// TIA Portal project "management parcare auto" (V17)

(* hardware
DEVICE "S7-1500/ET200MP station_1"  S7-1500 station
   slot 0: "Rail_0"  Rack  6ES7 590-1***0-0AA0
   slot 1: "PLC_1"  CPU 1511C-1 PN  6ES7 511-1CK01-0AB0  V2.5
      slot 3: "CPU display_1"  6ES7591-1AA00-0AA0
      slot 32768: "PROFINET interface_1"  X1
         slot 32769: "Port_1"  X1 P1
         slot 32770: "Port_2"  X1 P2
DEVICE "PC-System_1"  SIMATIC PC station
   slot 0: "SIMATIC PC station"  Rail  SIMATIC PC-Station  V1.0
      slot 125: "Stationmanager"  Station_Manager  V6.0.4
   slot 1: "HMI_RT_1"  WinCC RT Advanced  6AV2 104-0xxxx-xxxx  17.0.0.0
      slot 33792: "Computer interface"  Host interface
   slot 2: "CP 1628_1"  CP 1628  6GK1 162-8AA00  V8.2.2
DEVICE "HMI_1"  KTP700 Basic PN
   slot 0: "HMI_1"  KTP700 Basic PN  6AV2 123-2GB03-0AX0  15.1.0.0
   slot 1: "HMI_RT_2"  KTP700 Basic PN  6AV2 123-2GB03-0AX0  15.1.0.0
   slot 5: "HMI_1.IE_CP_1"  PROFINET Interface  15.0.1.0
      slot 1: "PROFINET Interface_1"  PROFINET Interface
         slot 1: "Port_1"  Port
*)

// ===== PLC "PLC_1"  CPU 1511C-1 PN =====

VAR_GLOBAL   // PLC tag table "Default tag table"
   "Exit barrier" AT %Q0.1 : Bool;
   "Entry barrier" AT %Q0.0 : Bool;
   "Entry sensor" AT %I0.0 : Bool;   // senzor bariera INTRARE
   "Exit sensor" AT %I1.0 : Bool;   // senzor barierea iesire
   "Parking lot 1 sensor" AT %I0.1 : Bool;   // senzor loc 1 (1-ocupat/ 0-liber)
   "Parking lot 2 sensor" AT %I0.2 : Bool;   // senzor loc 2
   "Parking lot 3 sensor" AT %I0.3 : Bool;
   "Parking lot 4 sensor" AT %I0.4 : Bool;
   "Parking lot 5 sensor" AT %I0.5 : Bool;
   "Parking lot 6 sensor" AT %I0.6 : Bool;
   "Parking lot 7 sensor" AT %I0.7 : Bool;
   "Parking lot 8 sensor" AT %I1.1 : Bool;
   "Parking lot 9 sensor" AT %I1.2 : Bool;
   "Parking lot 10 sensor" AT %I1.3 : Bool;
   "Number of cars" AT %MW20 : Int;   // nr de masini folosit la counter
   "System_Byte" AT %MB1 : Byte;
   "FirstScan" AT %M1.0 : Bool;
   "DiagStatusUpdate" AT %M1.1 : Bool;
   "AlwaysTRUE" AT %M1.2 : Bool;
   "AlwaysFALSE" AT %M1.3 : Bool;
   "Clock_Byte" AT %MB0 : Byte;
   "Clock_10Hz" AT %M0.0 : Bool;
   "Clock_5Hz" AT %M0.1 : Bool;
   "Clock_2.5Hz" AT %M0.2 : Bool;
   "Clock_2Hz" AT %M0.3 : Bool;
   "Clock_1.25Hz" AT %M0.4 : Bool;
   "Clock_1Hz" AT %M0.5 : Bool;
   "Clock_0.625Hz" AT %M0.6 : Bool;
   "Clock_0.5Hz" AT %M0.7 : Bool;
   "RdyToLog" AT %M2.0 : Bool;   // tagg folosit ca trigger pentru a rula vbScriptul
   "Tag5" AT %MW2 : Int;   // tagg folosit pentru counter pt animatie bariera intrare
   "Tag6" AT %MW4 : Int;   // tagg folosit pentru counter pt animatie bariera iesire
   "Tag_1" AT %M5.0 : Bool;
   "RdyToUpdate" AT %M6.0 : Bool;   // tagg folosit ca trigger pentru a rula vbSriptul de edit database
   "RdyToDelete" AT %M6.1 : Bool;   // tagg folosit ca trigger pentru a rula VbScriptul de stergere
   "Tag_2" AT %M6.2 : Bool;
   "Tag_3" AT %M6.3 : Bool;
   "Tag_4" AT %M6.4 : Bool;
   "Tag_5" AT %M6.5 : Bool;
   "Tag_6" AT %M6.6 : Bool;
   "Tag_7" AT %M6.7 : Bool;
   "Tag_8" AT %M5.1 : Bool;
   "Tag_9" AT %M5.2 : Bool;
   "Tag_10" AT %M5.3 : Bool;
   "Tag_11" AT %M5.4 : Bool;
   "Tag_12" AT %M7.0 : Bool;
   "Tag_13" AT %M7.1 : Bool;
   "Tag_14" AT %M7.2 : Bool;
   "Tag_15" AT %M7.3 : Bool;
   "Tag_16" AT %M7.4 : Bool;
   "Tag_17" AT %M7.5 : Bool;
   "Tag_18" AT %M7.6 : Bool;
   "Tag_19" AT %M7.7 : Bool;
   "Tag_20" AT %M8.0 : Bool;
   "Tag_21" AT %M8.1 : Bool;
END_VAR

// folder: DB's

DATA_BLOCK "02_DB_HMI_Buttons"   // DB2
{ S7_Optimized_Access := 'TRUE' }
VERSION : 0.1
   VAR
      pay : Bool;   // buton care simuleaza plata pentru a iesi din parcare
      "Parking lot 1" : Bool;   // buton in Hmi pentru a alege ce loc de parcare sa fie ocupat
      "Parking lot 2" : Bool;   // buton in Hmi pentru a alege ce loc de parcare sa fie ocupat
      "Parking lot 3" : Bool;   // buton in Hmi pentru a alege ce loc de parcare sa fie ocupat
      "Parking lot 4" : Bool;   // buton in Hmi pentru a alege ce loc de parcare sa fie ocupat
      "Parking lot 5" : Bool;   // buton in Hmi pentru a alege ce loc de parcare sa fie ocupat
      "Parking lot 6" : Bool;   // buton in Hmi pentru a alege ce loc de parcare sa fie ocupat
      "Parking lot 7" : Bool;   // buton in Hmi pentru a alege ce loc de parcare sa fie ocupat
      "Parking lot 8" : Bool;   // buton in Hmi pentru a alege ce loc de parcare sa fie ocupat
      "Parking lot 9" : Bool;   // buton in Hmi pentru a alege ce loc de parcare sa fie ocupat
      "Parking lot 10" : Bool;   // buton in Hmi pentru a alege ce loc de parcare sa fie ocupat
      "Entry button" : Bool;   // buton care simuleaza senzorul de intrare de la bariera
      "Exit button" : Bool;   // buton care simuleaza senzordul de iesire de la bariera
   END_VAR
   VAR RETAIN
      nrMasina_intrare : String;
   END_VAR
   VAR
      blank : String;
      nrMasina_iesire : String;
   END_VAR
BEGIN
END_DATA_BLOCK

DATA_BLOCK "04_DB_MarkersAuto"   // DB4
{ S7_Optimized_Access := 'TRUE' }
VERSION : 0.1
   VAR
      "car status_1" : Bool;
      "car status_2" : Bool;
      "car status_3" : Bool;
      "car status_4" : Bool;
      "car status_5" : Bool;
      "car status_6" : Bool;
      "car status_7" : Bool;
      "car status_8" : Bool;
      "car status_9" : Bool;
      "car status_10" : Bool;
      "remaining parking lots" : Int := 10;
      CarNumber : Int;   // dupa ce se introd un nr de masina, se face 1 , adica nr de masina a fost memorat
      "car status" : Bool;
      "Parking_lot_occupied 1" : Bool;   // locul a fost ocupat
      "Parking_lot_occupied 2" : Bool;
      "Parking_lot_occupied 3" : Bool;
      "Parking_lot_occupied 4" : Bool;
      "Parking_lot_occupied 5" : Bool;
      "Parking_lot_occupied 6" : Bool;
      "Parking_lot_occupied 7" : Bool;
      "Parking_lot_occupied 8" : Bool;
      "Parking_lot_occupied 9" : Bool;
      "Parking_lot_occupied 10" : Bool;
   END_VAR
BEGIN
END_DATA_BLOCK

DATA_BLOCK "05_DB_WinCC_buttons"   // DB5
{ S7_Optimized_Access := 'TRUE' }
VERSION : 0.1
   VAR
      loc_parcare_1 : Bool;   // buton de optiune pentru a alege locul de parcare 1
      loc_parcare_2 : Bool;   // -----//-------
      loc_parcare_3 : Bool;   // -----//-------
      loc_parcare_4 : Bool;   // -----//-------
      loc_parcare_5 : Bool;   // -----//-------
      loc_parcare_6 : Bool;   // -----//-------
      loc_parcare_7 : Bool;   // -----//-------
      loc_parcare_8 : Bool;   // -----//-------
      loc_parcare_9 : Bool;   // -----//-------
      loc_parcare_10 : Bool;   // -----//-------
      led_loc_1 : Bool;   // led pentru indicare loc de parcare( 1- rosu/ocupat; 0-verde/liber)
      led_loc_2 : Bool;   // led pentru indicare loc de parcare( 1- rosu/ocupat; 0-verde/liber)
      led_loc_3 : Bool;   // led pentru indicare loc de parcare( 1- rosu/ocupat; 0-verde/liber)
      led_loc_4 : Bool;   // led pentru indicare loc de parcare( 1- rosu/ocupat; 0-verde/liber)
      led_loc_5 : Bool;   // led pentru indicare loc de parcare( 1- rosu/ocupat; 0-verde/liber)
      led_loc_6 : Bool;   // led pentru indicare loc de parcare( 1- rosu/ocupat; 0-verde/liber)
      led_loc_7 : Bool;   // led pentru indicare loc de parcare( 1- rosu/ocupat; 0-verde/liber)
      led_loc_8 : Bool;   // led pentru indicare loc de parcare( 1- rosu/ocupat; 0-verde/liber)
      led_loc_9 : Bool;   // led pentru indicare loc de parcare( 1- rosu/ocupat; 0-verde/liber)
      led_loc_10 : Bool;   // led pentru indicare loc de parcare( 1- rosu/ocupat; 0-verde/liber)
      ResetNumber : Bool;
      ONBarrier_button_Entry : Bool;
      ONBarrier_button_Exit : Bool;
   END_VAR
BEGIN
END_DATA_BLOCK

DATA_BLOCK "01_FB_Setting_parameters_DB"   // DB6
{ S7_Optimized_Access := 'TRUE' }
VERSION : 0.1
// stored: InstanceOfName 01_FB_Setting_parameters
"01_FB_Setting_parameters"
BEGIN
END_DATA_BLOCK

DATA_BLOCK "08_DB_Alarms"   // DB8
{ S7_Optimized_Access := 'TRUE' }
VERSION : 0.1
   VAR
      Full : Word;   // Nu sunt locuri libere in parcare!
      Parking_lot_empty : Word;   // S-a intrat in parcare dar nu s-a ocupat niciun loc!
      EntryBarrierNotWorking : Word;   // Bariera de la intrare nu merge!
      ExitBarrierNotWorking : Word;   // Bariera de la iesire nu merge!
   END_VAR
BEGIN
END_DATA_BLOCK

DATA_BLOCK "11_DB_Inputs"   // DB11
{ S7_Optimized_Access := 'TRUE' }
VERSION : 0.1
   VAR
      "i0.0" : Bool;   // entry sensor / Senzor intrare
      "i0.1" : Bool;   // lot1
      "i0.2" : Bool;   // lot2
      "i0.3" : Bool;   // lot3
      "i0.4" : Bool;   // lot4
      "i0.5" : Bool;   // lot5
      "i0.6" : Bool;   // lot6
      "i0.7" : Bool;   // lot7
      "i1.0" : Bool;   // exit sensor / Senzor iesire
      "i1.1" : Bool;   // lot8
      "i1.2" : Bool;   // lot9
      "i1.3" : Bool;   // lot10
   END_VAR
BEGIN
END_DATA_BLOCK

// folder: Fc's

DATA_BLOCK "01_FB_Setting_parameters_DB_1"   // DB12
{ S7_Optimized_Access := 'TRUE' }
VERSION : 0.1
// stored: InstanceOfName 01_FB_Setting_parameters
"01_FB_Setting_parameters"
BEGIN
END_DATA_BLOCK

DATA_BLOCK "01_FB_Setting_parameters_DB_2"   // DB13
{ S7_Optimized_Access := 'TRUE' }
VERSION : 0.1
// stored: InstanceOfName 01_FB_Setting_parameters
"01_FB_Setting_parameters"
BEGIN
END_DATA_BLOCK

DATA_BLOCK "02_FB_exitLogic_DB_2"   // DB14
{ S7_Optimized_Access := 'TRUE' }
VERSION : 0.1
// stored: InstanceOfName 02_FB_exitLogic
"02_FB_exitLogic"
BEGIN
END_DATA_BLOCK

DATA_BLOCK "03_FB_entryLogic_DB"   // DB15
{ S7_Optimized_Access := 'TRUE' }
VERSION : 0.1
// stored: InstanceOfName 03_FB_entryLogic
"03_FB_entryLogic"
BEGIN
END_DATA_BLOCK

// folder: System blocks/Program resources

DATA_BLOCK "Client interface_1_Configuration"   // DB1
{ S7_Optimized_Access := 'TRUE' }
   VAR
      Connection : Struct
         ConnectInfo : OPC_UA_SessionConnectInfo;
         ConnectionHdl : DWord;
         ServerEndpointUrl : String[254];
      END_STRUCT;
      Namespaces : Struct
         NamespaceURIs : Array[0..0] of WString;
         ServerNamespaceIndexes : Array[0..0] of UInt;
         NamespaceStatusList : Array[0..0] of DWord;
         NamespaceCount : UInt;
      END_STRUCT;
      ReadLists : Struct
         "Read list_1" : Struct
            NodeCount : UInt;
            Nodes : Array[0..0] of OPC_UA_NodeId;
            NodeHdls : Array[0..0] of DWord;
         END_STRUCT;
      END_STRUCT;
   END_VAR
BEGIN
END_DATA_BLOCK

DATA_BLOCK "IEC_Counter_0_DB_1"   // DB7
{ S7_Optimized_Access := 'TRUE' }
AUTHOR : Simatic
FAMILY : IEC
NAME : CNTR
VERSION : 1.0
// stored: InstanceOfName IEC_COUNTER
"IEC_COUNTER"
BEGIN
END_DATA_BLOCK

DATA_BLOCK "IEC_Timer_0_DB_1"   // DB10
{ S7_Optimized_Access := 'TRUE' }
AUTHOR : Simatic
FAMILY : IEC
NAME : IEC_TMR
VERSION : 1.0
// stored: InstanceOfName IEC_TIMER
"IEC_TIMER"
BEGIN
END_DATA_BLOCK

// folder: (top level)

ORGANIZATION_BLOCK "Main"   // OB1, LAD, ProgramCycle
TITLE = "Main Program Sweep (Cycle)"
{ S7_Optimized_Access := 'TRUE' }
VERSION : 0.1
   VAR_INPUT
      Initial_Call : Bool;   // Initial call of this OB
      Remanence : Bool;   // =True, if remanent data are available
   END_VAR
BEGIN

REGION Network 1
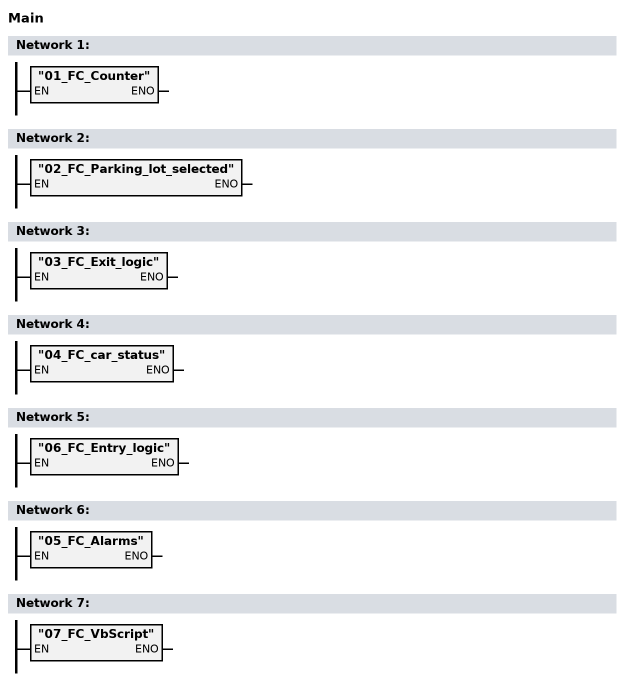
   RUNG wire#powerrail
      "01_FC_Counter"()
   END_RUNG
   // the same network as SCL:
   "01_FC_Counter"();
END_REGION

REGION Network 2
   RUNG wire#powerrail
      "02_FC_Parking_lot_selected"()
   END_RUNG
   // the same network as SCL:
   "02_FC_Parking_lot_selected"();
END_REGION

REGION Network 3
   RUNG wire#powerrail
      "03_FC_Exit_logic"()
   END_RUNG
   // the same network as SCL:
   "03_FC_Exit_logic"();
END_REGION

REGION Network 4
   RUNG wire#powerrail
      "04_FC_car_status"()
   END_RUNG
   // the same network as SCL:
   "04_FC_car_status"();
END_REGION

REGION Network 5
   RUNG wire#powerrail
      "06_FC_Entry_logic"()
   END_RUNG
   // the same network as SCL:
   "06_FC_Entry_logic"();
END_REGION

REGION Network 6
   RUNG wire#powerrail
      "05_FC_Alarms"()
   END_RUNG
   // the same network as SCL:
   "05_FC_Alarms"();
END_REGION

REGION Network 7
   RUNG wire#powerrail
      "07_FC_VbScript"()
   END_RUNG
   // the same network as SCL:
   "07_FC_VbScript"();
END_REGION
END_ORGANIZATION_BLOCK

// folder: FB's

FUNCTION_BLOCK "01_FB_Setting_parameters"   // FB1, LAD
{ S7_Optimized_Access := 'TRUE' }
VERSION : 0.1
   VAR_INPUT
      parking_lot_sensor : Bool;
   END_VAR
   VAR_OUTPUT
      parking_lot_occupied : Bool;   // locul de parcare respectiv a fost ocupat
   END_VAR
BEGIN

REGION Network 1: setare parametri pt un loc ocupat
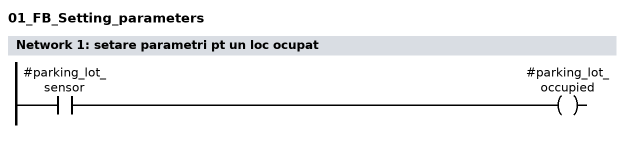
   RUNG wire#powerrail
      Contact( #parking_lot_sensor )
      Coil( #parking_lot_occupied )
   END_RUNG
   // the same network as SCL:
   #parking_lot_occupied := #parking_lot_sensor;
END_REGION
END_FUNCTION_BLOCK

FUNCTION_BLOCK "02_FB_exitLogic"   // FB2, LAD
{ S7_Optimized_Access := 'TRUE' }
VERSION : 0.1
   VAR_INPUT
      pay_button : Bool;
      "exit sensor" : Bool;
      manual : Bool;
   END_VAR
   VAR_OUTPUT
      barrier : Bool;
   END_VAR
BEGIN

REGION Network 1: logica iesire
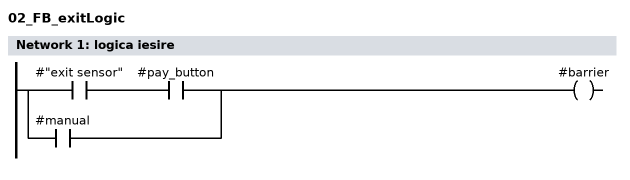
   RUNG wire#powerrail
      Contact( #"exit sensor" )
      Contact( #pay_button )
      wire#w1
      Coil( #barrier )
   END_RUNG
   RUNG wire#powerrail
      Contact( #manual )
   END_RUNG wire#w1
   // the same network as SCL:
   #barrier := (#"exit sensor" AND #pay_button) OR #manual;
END_REGION
END_FUNCTION_BLOCK

FUNCTION_BLOCK "03_FB_entryLogic"   // FB3, LAD
{ S7_Optimized_Access := 'TRUE' }
VERSION : 0.1
   VAR_INPUT
      entry_sensor : Bool;
      manual : Bool;
   END_VAR
   VAR_OUTPUT
      barrier : Bool;
   END_VAR
BEGIN

REGION Network 1
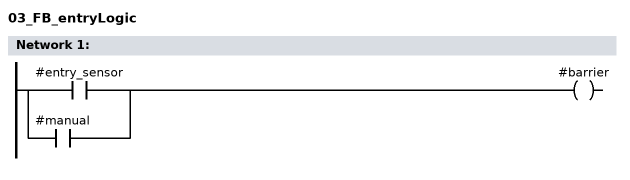
   RUNG wire#powerrail
      Contact( #entry_sensor )
      wire#w1
      Coil( #barrier )
   END_RUNG
   RUNG wire#powerrail
      Contact( #manual )
   END_RUNG wire#w1
   // the same network as SCL:
   #barrier := #entry_sensor OR #manual;
END_REGION
END_FUNCTION_BLOCK

// folder: Fc's

FUNCTION "01_FC_Counter" : Void   // FC1, LAD
{ S7_Optimized_Access := 'TRUE' }
VERSION : 0.1
   VAR CONSTANT
      i : Int := 1;
   END_VAR
   VAR_TEMP   // added for the SCL form of the ladder/FBD networks
      _w1 : Bool;
      _w2 : Bool;
      _w3 : Bool;
      _w4 : Bool;
      _w5 : Bool;
      _w6 : Bool;
      _w7 : Bool;
      _w8 : Bool;
      _w9 : Bool;
      _w10 : Bool;
   END_VAR
BEGIN

REGION Network 1: numar locuri ocupate
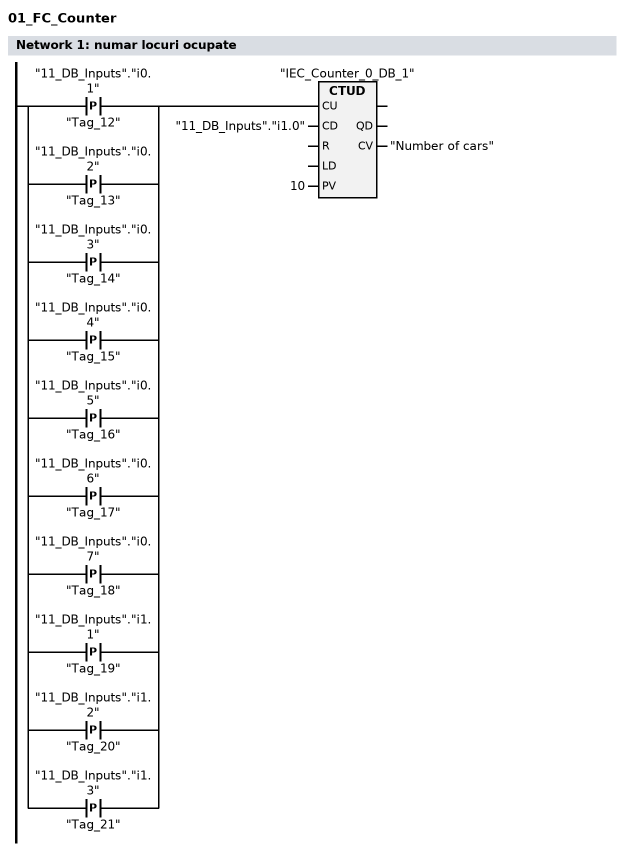
   #_w1 := "11_DB_Inputs"."i0.1" AND NOT "Tag_12";   // rising edge of "11_DB_Inputs"."i0.1"
   "Tag_12" := "11_DB_Inputs"."i0.1";
   #_w2 := "11_DB_Inputs"."i0.2" AND NOT "Tag_13";   // rising edge of "11_DB_Inputs"."i0.2"
   "Tag_13" := "11_DB_Inputs"."i0.2";
   #_w3 := "11_DB_Inputs"."i0.3" AND NOT "Tag_14";   // rising edge of "11_DB_Inputs"."i0.3"
   "Tag_14" := "11_DB_Inputs"."i0.3";
   #_w4 := "11_DB_Inputs"."i0.4" AND NOT "Tag_15";   // rising edge of "11_DB_Inputs"."i0.4"
   "Tag_15" := "11_DB_Inputs"."i0.4";
   #_w5 := "11_DB_Inputs"."i0.5" AND NOT "Tag_16";   // rising edge of "11_DB_Inputs"."i0.5"
   "Tag_16" := "11_DB_Inputs"."i0.5";
   #_w6 := "11_DB_Inputs"."i0.6" AND NOT "Tag_17";   // rising edge of "11_DB_Inputs"."i0.6"
   "Tag_17" := "11_DB_Inputs"."i0.6";
   #_w7 := "11_DB_Inputs"."i0.7" AND NOT "Tag_18";   // rising edge of "11_DB_Inputs"."i0.7"
   "Tag_18" := "11_DB_Inputs"."i0.7";
   #_w8 := "11_DB_Inputs"."i1.1" AND NOT "Tag_19";   // rising edge of "11_DB_Inputs"."i1.1"
   "Tag_19" := "11_DB_Inputs"."i1.1";
   #_w9 := "11_DB_Inputs"."i1.2" AND NOT "Tag_20";   // rising edge of "11_DB_Inputs"."i1.2"
   "Tag_20" := "11_DB_Inputs"."i1.2";
   #_w10 := "11_DB_Inputs"."i1.3" AND NOT "Tag_21";   // rising edge of "11_DB_Inputs"."i1.3"
   "Tag_21" := "11_DB_Inputs"."i1.3";
   "IEC_Counter_0_DB_1".CTUD(CU := #_w1 OR #_w2 OR #_w3 OR #_w4 OR #_w5 OR #_w6 OR #_w7 OR #_w8 OR #_w9 OR #_w10,
                           CD := "11_DB_Inputs"."i1.0",
                           PV := 10,
                           CV => "Number of cars");
END_REGION

REGION Network 2 (SCL): numar locuri libere

       "04_DB_MarkersAuto"."remaining parking lots" := 10 - "Number of cars";
END_REGION
END_FUNCTION

FUNCTION "02_FC_Parking_lot_selected" : Void   // FC2, LAD
{ S7_Optimized_Access := 'TRUE' }
VERSION : 0.1
BEGIN

REGION Network 1: loc 1 de parcare selectat
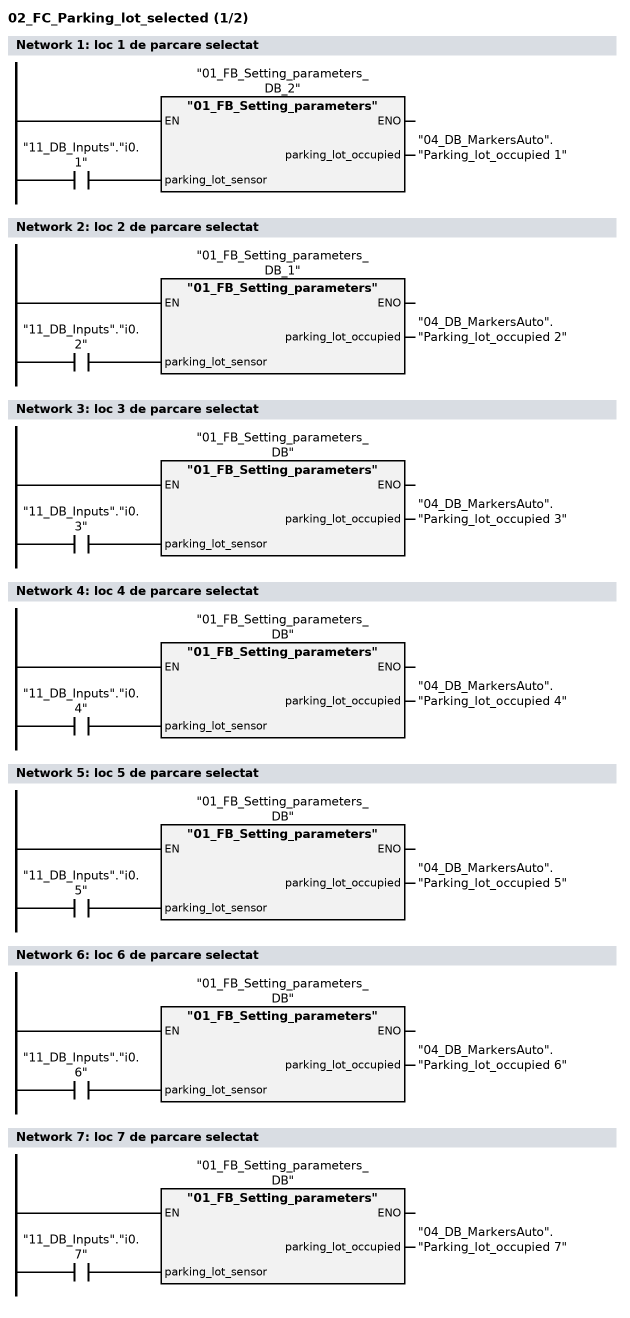
   RUNG wire#powerrail
      "01_FB_Setting_parameters_DB_2"(parking_lot_sensor := wire#w1, parking_lot_occupied => "04_DB_MarkersAuto"."Parking_lot_occupied 1")
   END_RUNG
   RUNG wire#powerrail
      Contact( "11_DB_Inputs"."i0.1" )
   END_RUNG wire#w1
   // the same network as SCL:
   "01_FB_Setting_parameters_DB_2"(parking_lot_sensor := "11_DB_Inputs"."i0.1",   // "01_FB_Setting_parameters"
                           parking_lot_occupied => "04_DB_MarkersAuto"."Parking_lot_occupied 1");
END_REGION

REGION Network 2: loc 2 de parcare selectat
   RUNG wire#powerrail
      "01_FB_Setting_parameters_DB_1"(parking_lot_sensor := wire#w1, parking_lot_occupied => "04_DB_MarkersAuto"."Parking_lot_occupied 2")
   END_RUNG
   RUNG wire#powerrail
      Contact( "11_DB_Inputs"."i0.2" )
   END_RUNG wire#w1
   // the same network as SCL:
   "01_FB_Setting_parameters_DB_1"(parking_lot_sensor := "11_DB_Inputs"."i0.2",   // "01_FB_Setting_parameters"
                           parking_lot_occupied => "04_DB_MarkersAuto"."Parking_lot_occupied 2");
END_REGION

REGION Network 3: loc 3 de parcare selectat
   RUNG wire#powerrail
      "01_FB_Setting_parameters_DB"(parking_lot_sensor := wire#w1, parking_lot_occupied => "04_DB_MarkersAuto"."Parking_lot_occupied 3")
   END_RUNG
   RUNG wire#powerrail
      Contact( "11_DB_Inputs"."i0.3" )
   END_RUNG wire#w1
   // the same network as SCL:
   "01_FB_Setting_parameters_DB"(parking_lot_sensor := "11_DB_Inputs"."i0.3",   // "01_FB_Setting_parameters"
                           parking_lot_occupied => "04_DB_MarkersAuto"."Parking_lot_occupied 3");
END_REGION

REGION Network 4: loc 4 de parcare selectat
   RUNG wire#powerrail
      "01_FB_Setting_parameters_DB"(parking_lot_sensor := wire#w1, parking_lot_occupied => "04_DB_MarkersAuto"."Parking_lot_occupied 4")
   END_RUNG
   RUNG wire#powerrail
      Contact( "11_DB_Inputs"."i0.4" )
   END_RUNG wire#w1
   // the same network as SCL:
   "01_FB_Setting_parameters_DB"(parking_lot_sensor := "11_DB_Inputs"."i0.4",   // "01_FB_Setting_parameters"
                           parking_lot_occupied => "04_DB_MarkersAuto"."Parking_lot_occupied 4");
END_REGION

REGION Network 5: loc 5 de parcare selectat
   RUNG wire#powerrail
      "01_FB_Setting_parameters_DB"(parking_lot_sensor := wire#w1, parking_lot_occupied => "04_DB_MarkersAuto"."Parking_lot_occupied 5")
   END_RUNG
   RUNG wire#powerrail
      Contact( "11_DB_Inputs"."i0.5" )
   END_RUNG wire#w1
   // the same network as SCL:
   "01_FB_Setting_parameters_DB"(parking_lot_sensor := "11_DB_Inputs"."i0.5",   // "01_FB_Setting_parameters"
                           parking_lot_occupied => "04_DB_MarkersAuto"."Parking_lot_occupied 5");
END_REGION

REGION Network 6: loc 6 de parcare selectat
   RUNG wire#powerrail
      "01_FB_Setting_parameters_DB"(parking_lot_sensor := wire#w1, parking_lot_occupied => "04_DB_MarkersAuto"."Parking_lot_occupied 6")
   END_RUNG
   RUNG wire#powerrail
      Contact( "11_DB_Inputs"."i0.6" )
   END_RUNG wire#w1
   // the same network as SCL:
   "01_FB_Setting_parameters_DB"(parking_lot_sensor := "11_DB_Inputs"."i0.6",   // "01_FB_Setting_parameters"
                           parking_lot_occupied => "04_DB_MarkersAuto"."Parking_lot_occupied 6");
END_REGION

REGION Network 7: loc 7 de parcare selectat
   RUNG wire#powerrail
      "01_FB_Setting_parameters_DB"(parking_lot_sensor := wire#w1, parking_lot_occupied => "04_DB_MarkersAuto"."Parking_lot_occupied 7")
   END_RUNG
   RUNG wire#powerrail
      Contact( "11_DB_Inputs"."i0.7" )
   END_RUNG wire#w1
   // the same network as SCL:
   "01_FB_Setting_parameters_DB"(parking_lot_sensor := "11_DB_Inputs"."i0.7",   // "01_FB_Setting_parameters"
                           parking_lot_occupied => "04_DB_MarkersAuto"."Parking_lot_occupied 7");
END_REGION

REGION Network 8: loc 8 de parcare selectat
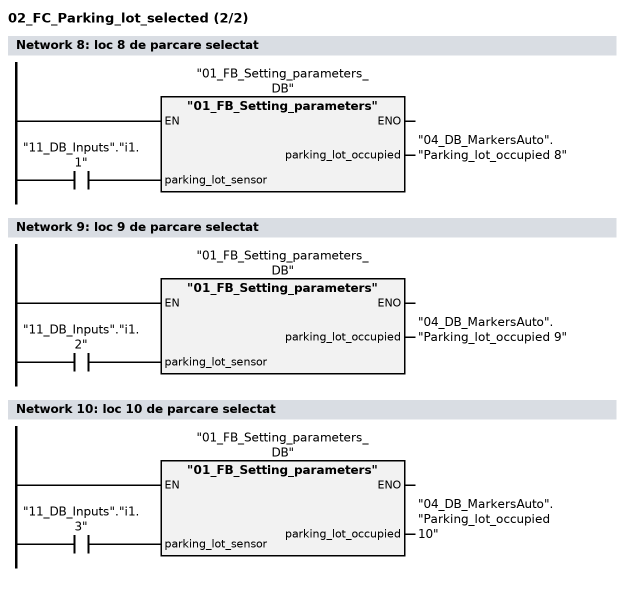
   RUNG wire#powerrail
      "01_FB_Setting_parameters_DB"(parking_lot_sensor := wire#w1, parking_lot_occupied => "04_DB_MarkersAuto"."Parking_lot_occupied 8")
   END_RUNG
   RUNG wire#powerrail
      Contact( "11_DB_Inputs"."i1.1" )
   END_RUNG wire#w1
   // the same network as SCL:
   "01_FB_Setting_parameters_DB"(parking_lot_sensor := "11_DB_Inputs"."i1.1",   // "01_FB_Setting_parameters"
                           parking_lot_occupied => "04_DB_MarkersAuto"."Parking_lot_occupied 8");
END_REGION

REGION Network 9: loc 9 de parcare selectat
   RUNG wire#powerrail
      "01_FB_Setting_parameters_DB"(parking_lot_sensor := wire#w1, parking_lot_occupied => "04_DB_MarkersAuto"."Parking_lot_occupied 9")
   END_RUNG
   RUNG wire#powerrail
      Contact( "11_DB_Inputs"."i1.2" )
   END_RUNG wire#w1
   // the same network as SCL:
   "01_FB_Setting_parameters_DB"(parking_lot_sensor := "11_DB_Inputs"."i1.2",   // "01_FB_Setting_parameters"
                           parking_lot_occupied => "04_DB_MarkersAuto"."Parking_lot_occupied 9");
END_REGION

REGION Network 10: loc 10 de parcare selectat
   RUNG wire#powerrail
      "01_FB_Setting_parameters_DB"(parking_lot_sensor := wire#w1, parking_lot_occupied => "04_DB_MarkersAuto"."Parking_lot_occupied 10")
   END_RUNG
   RUNG wire#powerrail
      Contact( "11_DB_Inputs"."i1.3" )
   END_RUNG wire#w1
   // the same network as SCL:
   "01_FB_Setting_parameters_DB"(parking_lot_sensor := "11_DB_Inputs"."i1.3",   // "01_FB_Setting_parameters"
                           parking_lot_occupied => "04_DB_MarkersAuto"."Parking_lot_occupied 10");
END_REGION
END_FUNCTION

FUNCTION "03_FC_Exit_logic" : Void   // FC3, LAD
{ S7_Optimized_Access := 'TRUE' }
VERSION : 0.1
BEGIN

REGION Network 1
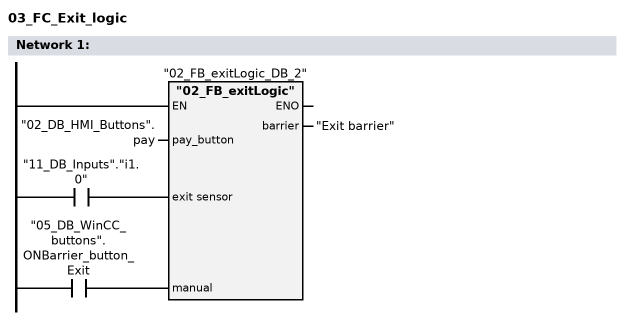
   RUNG wire#powerrail
      "02_FB_exitLogic_DB_2"("exit sensor" := wire#w1, manual := wire#w2, pay_button := "02_DB_HMI_Buttons".pay, barrier => "Exit barrier")
   END_RUNG
   RUNG wire#powerrail
      Contact( "11_DB_Inputs"."i1.0" )
   END_RUNG wire#w1
   RUNG wire#powerrail
      Contact( "05_DB_WinCC_buttons".ONBarrier_button_Exit )
   END_RUNG wire#w2
   // the same network as SCL:
   "02_FB_exitLogic_DB_2"(pay_button := "02_DB_HMI_Buttons".pay,   // "02_FB_exitLogic"
                          "exit sensor" := "11_DB_Inputs"."i1.0",
                          manual := "05_DB_WinCC_buttons".ONBarrier_button_Exit,
                          barrier => "Exit barrier");
END_REGION
END_FUNCTION

FUNCTION "04_FC_car_status" : Void   // FC4, LAD
{ S7_Optimized_Access := 'TRUE' }
VERSION : 0.1
BEGIN

REGION Network 1: stergere nr masina din I/O field dupa ce senzorul de intrare e zero
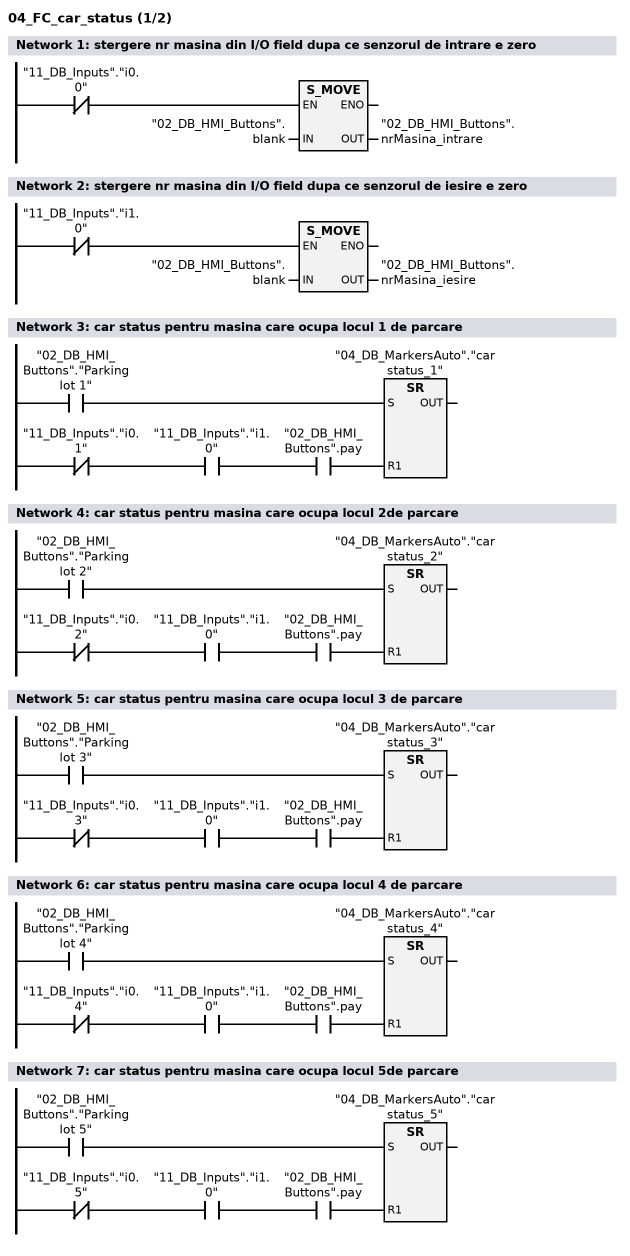
   RUNG wire#powerrail
      I_Contact( "11_DB_Inputs"."i0.0" )
      S_Move(in := "02_DB_HMI_Buttons".blank, out => "02_DB_HMI_Buttons".nrMasina_intrare)
   END_RUNG
   // the same network as SCL:
   IF NOT "11_DB_Inputs"."i0.0" THEN
       "02_DB_HMI_Buttons".nrMasina_intrare := "02_DB_HMI_Buttons".blank;
   END_IF;
END_REGION

REGION Network 2: stergere nr masina din I/O field dupa ce senzorul de iesire e zero
   RUNG wire#powerrail
      I_Contact( "11_DB_Inputs"."i1.0" )
      S_Move(in := "02_DB_HMI_Buttons".blank, out => "02_DB_HMI_Buttons".nrMasina_iesire)
   END_RUNG
   // the same network as SCL:
   IF NOT "11_DB_Inputs"."i1.0" THEN
       "02_DB_HMI_Buttons".nrMasina_iesire := "02_DB_HMI_Buttons".blank;
   END_IF;
END_REGION

REGION Network 3: car status pentru masina care ocupa locul 1 de parcare
   RUNG wire#powerrail
      Contact( "02_DB_HMI_Buttons"."Parking lot 1" )
      S_SR(operand := "04_DB_MarkersAuto"."car status_1", r1 := wire#w1)
   END_RUNG
   RUNG wire#powerrail
      I_Contact( "11_DB_Inputs"."i0.1" )
      Contact( "11_DB_Inputs"."i1.0" )
      Contact( "02_DB_HMI_Buttons".pay )
   END_RUNG wire#w1
   // the same network as SCL:
   IF "02_DB_HMI_Buttons"."Parking lot 1" THEN
       "04_DB_MarkersAuto"."car status_1" := TRUE;   // SR flip-flop
   END_IF;
   IF NOT "11_DB_Inputs"."i0.1" AND "11_DB_Inputs"."i1.0" AND "02_DB_HMI_Buttons".pay THEN
       "04_DB_MarkersAuto"."car status_1" := FALSE;
   END_IF;
END_REGION

REGION Network 4: car status pentru masina care ocupa locul 2de parcare
   RUNG wire#powerrail
      Contact( "02_DB_HMI_Buttons"."Parking lot 2" )
      S_SR(operand := "04_DB_MarkersAuto"."car status_2", r1 := wire#w1)
   END_RUNG
   RUNG wire#powerrail
      I_Contact( "11_DB_Inputs"."i0.2" )
      Contact( "11_DB_Inputs"."i1.0" )
      Contact( "02_DB_HMI_Buttons".pay )
   END_RUNG wire#w1
   // the same network as SCL:
   IF "02_DB_HMI_Buttons"."Parking lot 2" THEN
       "04_DB_MarkersAuto"."car status_2" := TRUE;   // SR flip-flop
   END_IF;
   IF NOT "11_DB_Inputs"."i0.2" AND "11_DB_Inputs"."i1.0" AND "02_DB_HMI_Buttons".pay THEN
       "04_DB_MarkersAuto"."car status_2" := FALSE;
   END_IF;
END_REGION

REGION Network 5: car status pentru masina care ocupa locul 3 de parcare
   RUNG wire#powerrail
      Contact( "02_DB_HMI_Buttons"."Parking lot 3" )
      S_SR(operand := "04_DB_MarkersAuto"."car status_3", r1 := wire#w1)
   END_RUNG
   RUNG wire#powerrail
      I_Contact( "11_DB_Inputs"."i0.3" )
      Contact( "11_DB_Inputs"."i1.0" )
      Contact( "02_DB_HMI_Buttons".pay )
   END_RUNG wire#w1
   // the same network as SCL:
   IF "02_DB_HMI_Buttons"."Parking lot 3" THEN
       "04_DB_MarkersAuto"."car status_3" := TRUE;   // SR flip-flop
   END_IF;
   IF NOT "11_DB_Inputs"."i0.3" AND "11_DB_Inputs"."i1.0" AND "02_DB_HMI_Buttons".pay THEN
       "04_DB_MarkersAuto"."car status_3" := FALSE;
   END_IF;
END_REGION

REGION Network 6: car status pentru masina care ocupa locul 4 de parcare
   RUNG wire#powerrail
      Contact( "02_DB_HMI_Buttons"."Parking lot 4" )
      S_SR(operand := "04_DB_MarkersAuto"."car status_4", r1 := wire#w1)
   END_RUNG
   RUNG wire#powerrail
      I_Contact( "11_DB_Inputs"."i0.4" )
      Contact( "11_DB_Inputs"."i1.0" )
      Contact( "02_DB_HMI_Buttons".pay )
   END_RUNG wire#w1
   // the same network as SCL:
   IF "02_DB_HMI_Buttons"."Parking lot 4" THEN
       "04_DB_MarkersAuto"."car status_4" := TRUE;   // SR flip-flop
   END_IF;
   IF NOT "11_DB_Inputs"."i0.4" AND "11_DB_Inputs"."i1.0" AND "02_DB_HMI_Buttons".pay THEN
       "04_DB_MarkersAuto"."car status_4" := FALSE;
   END_IF;
END_REGION

REGION Network 7: car status pentru masina care ocupa locul 5de parcare
   RUNG wire#powerrail
      Contact( "02_DB_HMI_Buttons"."Parking lot 5" )
      S_SR(operand := "04_DB_MarkersAuto"."car status_5", r1 := wire#w1)
   END_RUNG
   RUNG wire#powerrail
      I_Contact( "11_DB_Inputs"."i0.5" )
      Contact( "11_DB_Inputs"."i1.0" )
      Contact( "02_DB_HMI_Buttons".pay )
   END_RUNG wire#w1
   // the same network as SCL:
   IF "02_DB_HMI_Buttons"."Parking lot 5" THEN
       "04_DB_MarkersAuto"."car status_5" := TRUE;   // SR flip-flop
   END_IF;
   IF NOT "11_DB_Inputs"."i0.5" AND "11_DB_Inputs"."i1.0" AND "02_DB_HMI_Buttons".pay THEN
       "04_DB_MarkersAuto"."car status_5" := FALSE;
   END_IF;
END_REGION

REGION Network 8: car status pentru masina care ocupa locul 6 de parcare